(* Logix 5000 project; controller PLC_MCC1300_75F1 vendor 1 type 14 code 166 rev 32.11; software revision 32.04; part 55 of 83 *)
(* tags used below, declared in another part *)
   CM_AreaStackerToLine_JS1 : CM_AreaStackerToLine;
   CM_AreaStackerToLine_JS1_Sync : CM_AreaStackerToLine;
   CM_ConveyorStackerToLine_JS1_Sync : CM_ConveyorStackerToLine;
   Convoy_SL_DATA_NULL : UDT_Convoy_SL;
   GP_AccessArea_M311S_STC : GP_AccessArea_STC;
   GP_InvertCapxLite : GP_InvertCapxLite;
   GP_M311A : GP_Rotator;
   GP_OB_InitializeMain : GP_OB_Initialize;
   GP_ScadaPlate : GP_ScadaPlate;
   Gp_SpaceConvUtilities_V1 : GP_SpaceConvUtilities_V1;
   M310B : MAC_Conveyor;
   M310B_Data : UDT_Convoy_SL;
   M310B_SpaceConv_Utilities : SpaceConv_Utilities;
   M311 : MAC_Conveyor;
   M311_ALM : MAC_Conveyor_ALM;
   M311_Data : UDT_Convoy_SL;
   M311_dLastRotationA_ID : DINT;
   M311_HMR : MAC_Conveyor_HMR;
   M311_HMW : MAC_Conveyor_HMW;
   M311_M1_DR : AXIS_CIP_DRIVE;
   M311_M1_DR_IN_MAM : MOTION_INSTRUCTION;
   M311_SpaceConv_Utilities : SpaceConv_Utilities;
   M311_TON_Synchro_timeout : TIMER;
   M311_xOS_SentToCullet : BOOL;
   M311_xSendCulletReqActive : BOOL;
   M311_xSensorTimeout : BOOL;
   M311A : MAC_Rotator;
   M311A_Data : UDT_Convoy_SL;
   M311A_HMR : MAC_Rotator_HMR;
   M311A_HMW : MAC_Rotator_HMW;
   M311A_M1_DR : AXIS_CIP_DRIVE;
   M311A_M1_DR_IN_MAM : MOTION_INSTRUCTION;
   M311A_rLastPosition : REAL;
   M311M312_OffsetBaricentre_cmm : DINT;
   M312 : MAC_Conveyor_Single;
   M312_Data : UDT_Convoy_SL;
   M312_SpaceConv_Utilities : SpaceConv_Utilities;
   O : INT[128];
   Sbr_OUT_ReqRot_CW : BOOL;
   TMP_d : DINT;
   TMP_dActualOnLHS : DINT;
   TMP_dDecelerationPositionEndConveyor : DINT;
   TMP_dMissingOnLHS : DINT;
   TMP_dOffsetLoadUnload_cmm : DINT;
   TMP_HeadPos : DINT;
   TMP_Portrait : BOOL;
   TMP_SendToCullet : BOOL;
   TMP_x : BOOL;
   TMP_xConveyorOfStartCleaning : BOOL;
   TMP_xEnableZoneCleaning : BOOL;
   TMP_xJustOnePlateMissing : BOOL;
   TMP_xLiteThisDestPresent : BOOL;
   x311PortraitMode : BOOL;
   xAlwaysOFF : BOOL;
   xAlwaysON : BOOL;
   xDebugOFF : BOOL;
   Z401 : MAC_Zone;
   Z401_HMI_rgtPlateScada_Internal : HMI_LiteData[5,2,7];
   Z401_HMR : MAC_Zone_HMR;
   Z401S_INPUT_xSafetyAreaPopup : BOOL;
(* MainProgram, continued *)

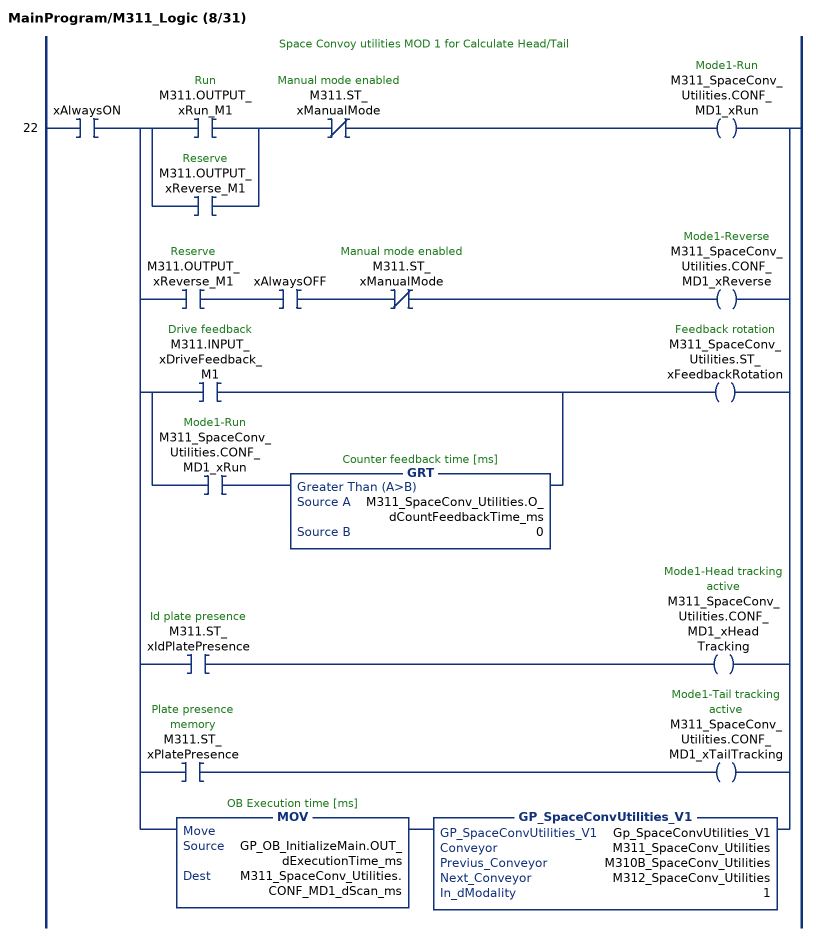
   [picture p890: MainProgram/M311_Logic rungs 22-22]
   // Space Convoy utilities MOD 1 for Calculate Head/Tail
   22: XIC(xAlwaysON)[[XIC(M311.OUTPUT_xRun_M1) ,XIC(M311.OUTPUT_xReverse_M1) ] XIO(M311.ST_xManualMode) OTE(M311_SpaceConv_Utilities.CONF_MD1_xRun) ,XIC(M311.OUTPUT_xReverse_M1) XIC(xAlwaysOFF) XIO(M311.ST_xManualMode) OTE(M311_SpaceConv_Utilities.CONF_MD1_xReverse) ,[XIC(M311.INPUT_xDriveFeedback_M1) ,XIC(M311_SpaceConv_Utilities.CONF_MD1_xRun) GRT(M311_SpaceConv_Utilities.O_dCountFeedbackTime_ms,0) ] OTE(M311_SpaceConv_Utilities.ST_xFeedbackRotation) ,XIC(M311.ST_xIdPlatePresence) OTE(M311_SpaceConv_Utilities.CONF_MD1_xHeadTracking) ,XIC(M311.ST_xPlatePresence) OTE(M311_SpaceConv_Utilities.CONF_MD1_xTailTracking) ,MOV(GP_OB_InitializeMain.OUT_dExecutionTime_ms,M311_SpaceConv_Utilities.CONF_MD1_dScan_ms) GP_SpaceConvUtilities_V1(Gp_SpaceConvUtilities_V1,M311_SpaceConv_Utilities,M310B_SpaceConv_Utilities,M312_SpaceConv_Utilities,1) ];
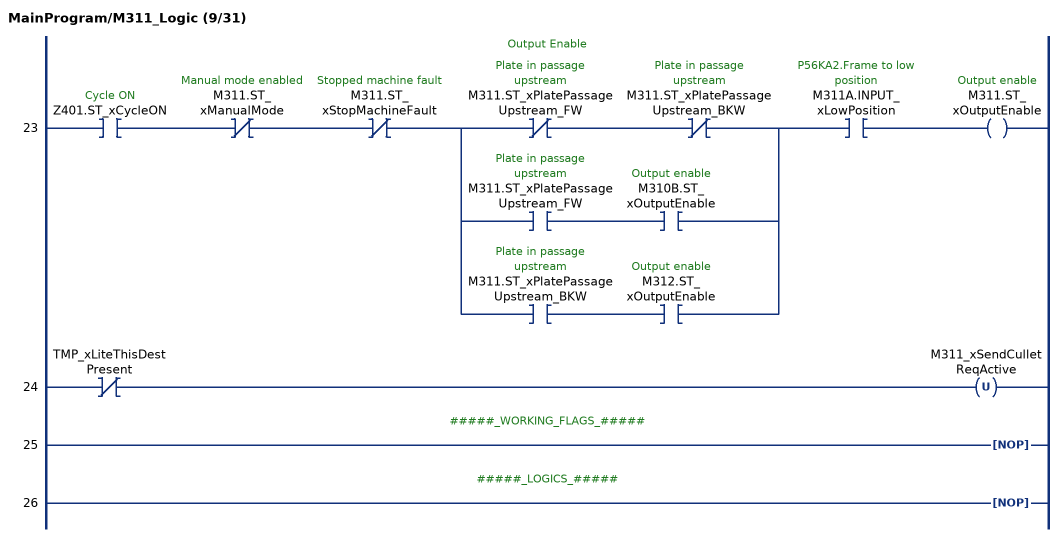
   // Output Enable
   23: XIC(Z401.ST_xCycleON)XIO(M311.ST_xManualMode)XIO(M311.ST_xStopMachineFault)[XIO(M311.ST_xPlatePassageUpstream_FW) XIO(M311.ST_xPlatePassageUpstream_BKW) ,XIC(M311.ST_xPlatePassageUpstream_FW) XIC(M310B.ST_xOutputEnable) ,XIC(M311.ST_xPlatePassageUpstream_BKW) XIC(M312.ST_xOutputEnable) ]XIC(M311A.INPUT_xLowPosition)OTE(M311.ST_xOutputEnable);
   24: XIO(TMP_xLiteThisDestPresent)OTU(M311_xSendCulletReqActive);
   // #####_WORKING_FLAGS_#####
   25: NOP();
   // #####_LOGICS_#####
   26: NOP();
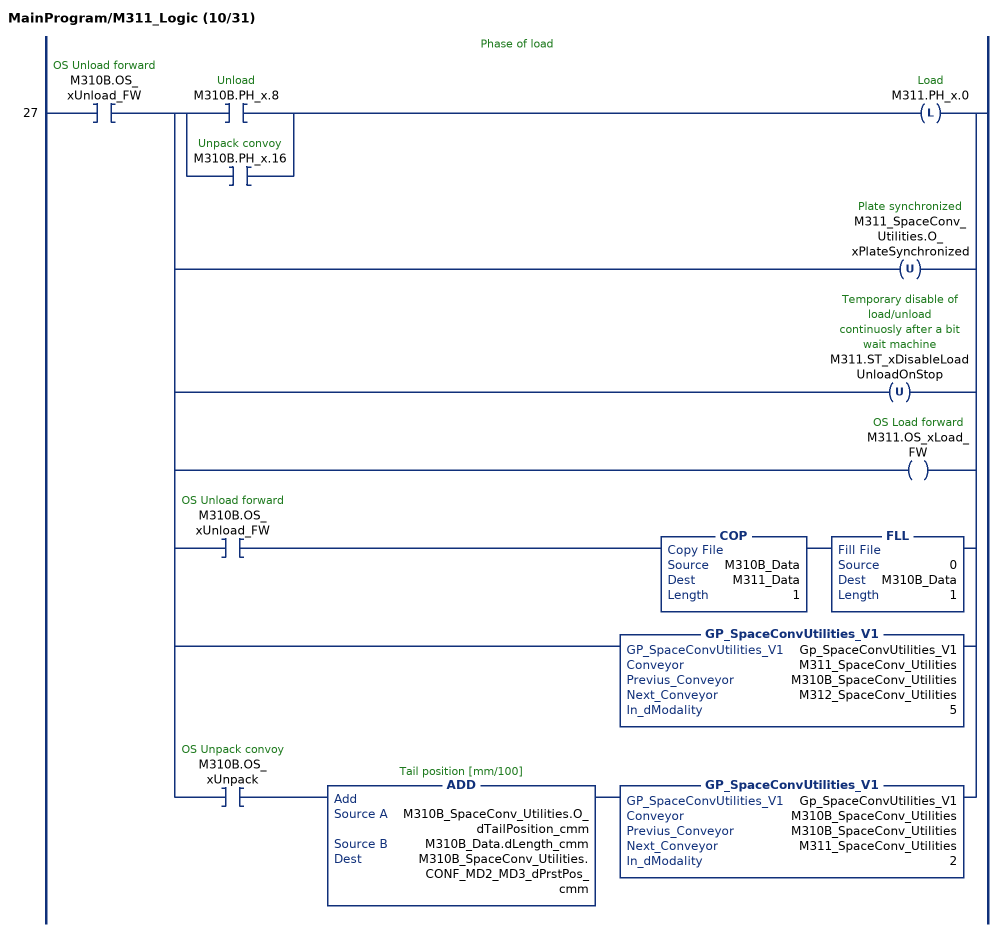
   // Phase of load
   27: XIC(M310B.OS_xUnload_FW)[[XIC(M310B.PH_x.8) ,XIC(M310B.PH_x.16) ] OTL(M311.PH_x.0) ,OTU(M311_SpaceConv_Utilities.O_xPlateSynchronized) ,OTU(M311.ST_xDisableLoadUnloadOnStop) ,OTE(M311.OS_xLoad_FW) ,XIC(M310B.OS_xUnload_FW) COP(M310B_Data,M311_Data,1) FLL(0,M310B_Data,1) ,GP_SpaceConvUtilities_V1(Gp_SpaceConvUtilities_V1,M311_SpaceConv_Utilities,M310B_SpaceConv_Utilities,M312_SpaceConv_Utilities,5) ,XIC(M310B.OS_xUnpack) ADD(M310B_SpaceConv_Utilities.O_dTailPosition_cmm,M310B_Data.dLength_cmm,M310B_SpaceConv_Utilities.CONF_MD2_MD3_dPrstPos_cmm) GP_SpaceConvUtilities_V1(Gp_SpaceConvUtilities_V1,M310B_SpaceConv_Utilities,M310B_SpaceConv_Utilities,M311_SpaceConv_Utilities,2) ];
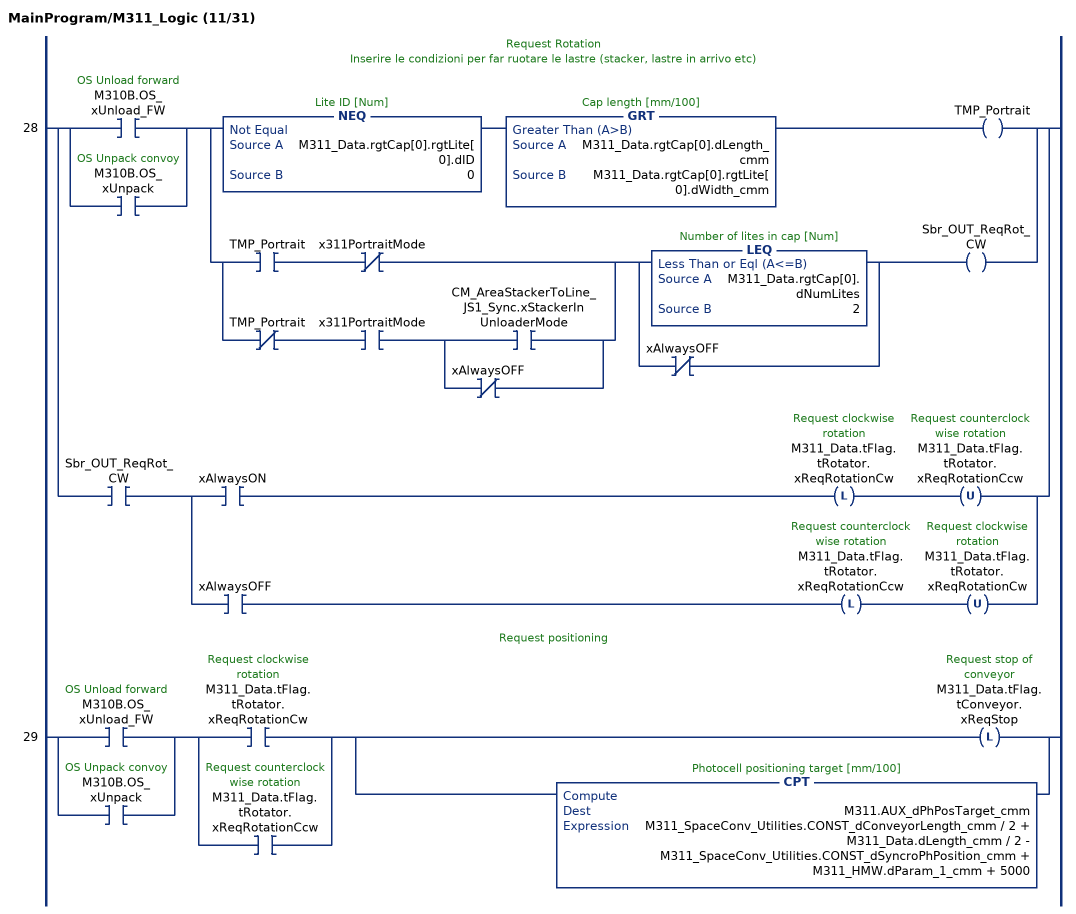
   // Request Rotation
   // Inserire le condizioni per far ruotare le lastre (stacker, lastre in arrivo etc)
   28: [[XIC(M310B.OS_xUnload_FW) ,XIC(M310B.OS_xUnpack) ] [NEQ(M311_Data.rgtCap[0].rgtLite[0].dID,0) GRT(M311_Data.rgtCap[0].dLength_cmm,M311_Data.rgtCap[0].rgtLite[0].dWidth_cmm) OTE(TMP_Portrait) ,[XIC(TMP_Portrait) XIO(x311PortraitMode) ,XIO(TMP_Portrait) XIC(x311PortraitMode) [XIC(CM_AreaStackerToLine_JS1_Sync.xStackerInUnloaderMode) ,XIO(xAlwaysOFF) ] ] [LEQ(M311_Data.rgtCap[0].dNumLites,2) ,XIO(xAlwaysOFF) ] OTE(Sbr_OUT_ReqRot_CW) ] ,XIC(Sbr_OUT_ReqRot_CW) [XIC(xAlwaysON) OTL(M311_Data.tFlag.tRotator.xReqRotationCw) OTU(M311_Data.tFlag.tRotator.xReqRotationCcw) ,XIC(xAlwaysOFF) OTL(M311_Data.tFlag.tRotator.xReqRotationCcw) OTU(M311_Data.tFlag.tRotator.xReqRotationCw) ] ];
   // Request positioning
   29: [XIC(M310B.OS_xUnload_FW) ,XIC(M310B.OS_xUnpack) ][XIC(M311_Data.tFlag.tRotator.xReqRotationCw) ,XIC(M311_Data.tFlag.tRotator.xReqRotationCcw) ][OTL(M311_Data.tFlag.tConveyor.xReqStop) ,CPT(M311.AUX_dPhPosTarget_cmm,M311_SpaceConv_Utilities.CONST_dConveyorLength_cmm / 2 + M311_Data.dLength_cmm / 2 - M311_SpaceConv_Utilities.CONST_dSyncroPhPosition_cmm + M311_HMW.dParam_1_cmm + 5000) ];
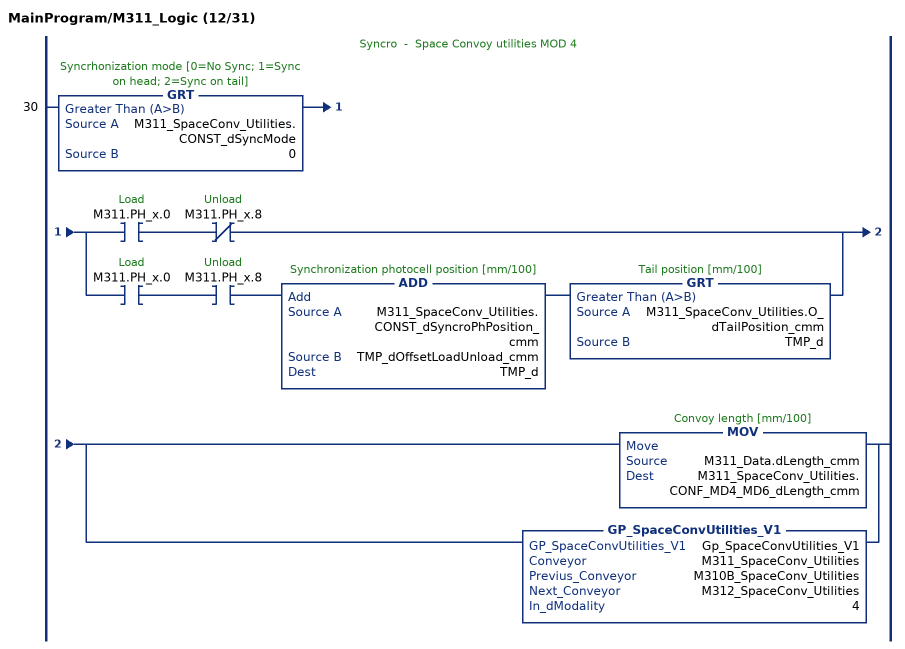
   // Syncro  -  Space Convoy utilities MOD 4
   30: GRT(M311_SpaceConv_Utilities.CONST_dSyncMode,0)[XIC(M311.PH_x.0) XIO(M311.PH_x.8) ,XIC(M311.PH_x.0) XIC(M311.PH_x.8) ADD(M311_SpaceConv_Utilities.CONST_dSyncroPhPosition_cmm,TMP_dOffsetLoadUnload_cmm,TMP_d) GRT(M311_SpaceConv_Utilities.O_dTailPosition_cmm,TMP_d) ][MOV(M311_Data.dLength_cmm,M311_SpaceConv_Utilities.CONF_MD4_MD6_dLength_cmm) ,GP_SpaceConvUtilities_V1(Gp_SpaceConvUtilities_V1,M311_SpaceConv_Utilities,M310B_SpaceConv_Utilities,M312_SpaceConv_Utilities,4) ];
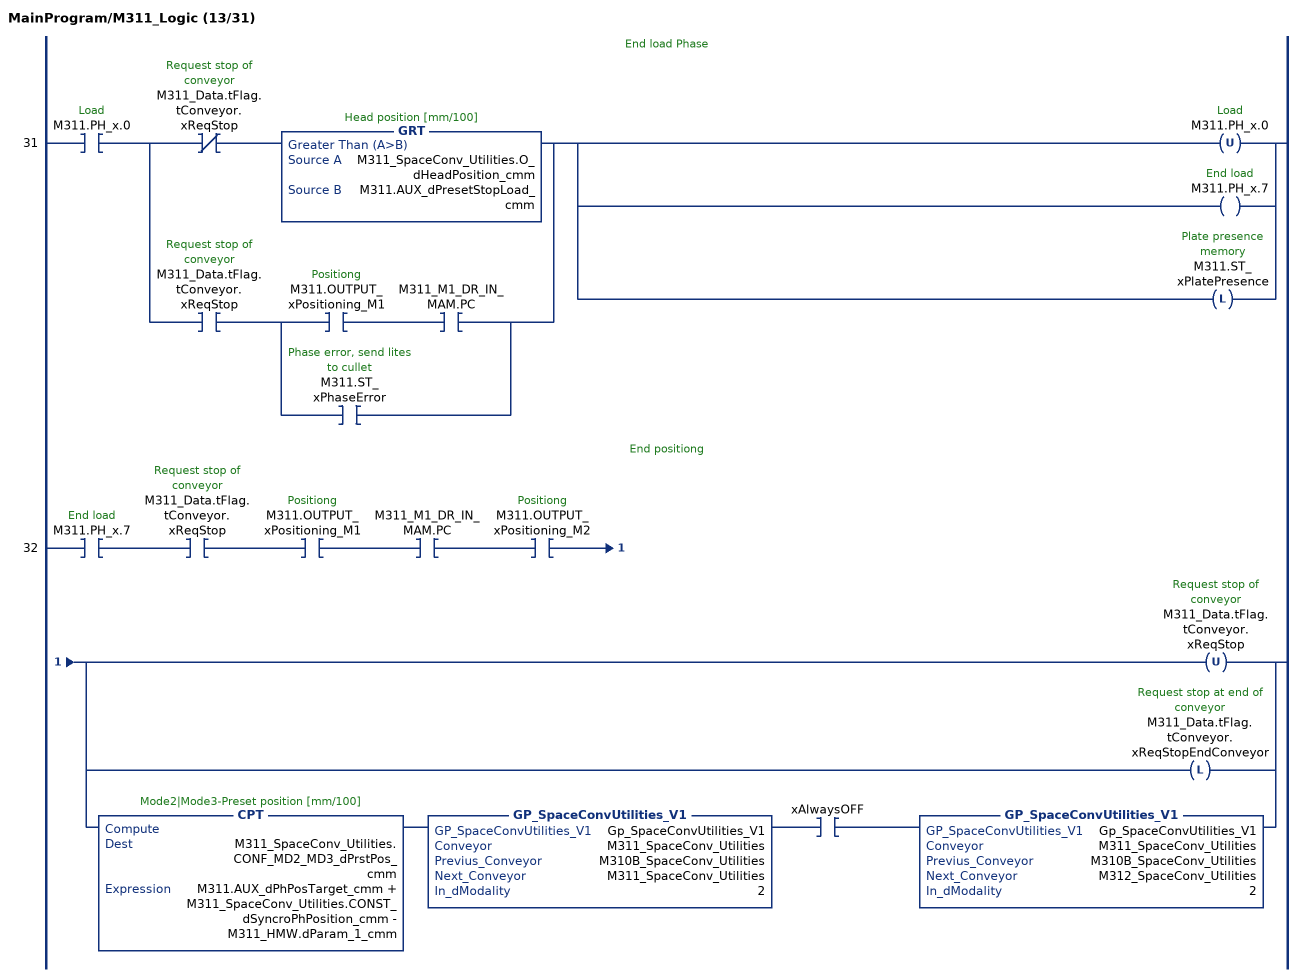
   // End load Phase
   31: XIC(M311.PH_x.0)[XIO(M311_Data.tFlag.tConveyor.xReqStop) GRT(M311_SpaceConv_Utilities.O_dHeadPosition_cmm,M311.AUX_dPresetStopLoad_cmm) ,XIC(M311_Data.tFlag.tConveyor.xReqStop) [XIC(M311.OUTPUT_xPositioning_M1) XIC(M311_M1_DR_IN_MAM.PC) ,XIC(M311.ST_xPhaseError) ] ][OTU(M311.PH_x.0) ,OTE(M311.PH_x.7) ,OTL(M311.ST_xPlatePresence) ];
   // End positiong
   32: XIC(M311.PH_x.7)XIC(M311_Data.tFlag.tConveyor.xReqStop)XIC(M311.OUTPUT_xPositioning_M1)XIC(M311_M1_DR_IN_MAM.PC)XIC(M311.OUTPUT_xPositioning_M2)[OTU(M311_Data.tFlag.tConveyor.xReqStop) ,OTL(M311_Data.tFlag.tConveyor.xReqStopEndConveyor) ,CPT(M311_SpaceConv_Utilities.CONF_MD2_MD3_dPrstPos_cmm,M311.AUX_dPhPosTarget_cmm + M311_SpaceConv_Utilities.CONST_dSyncroPhPosition_cmm - M311_HMW.dParam_1_cmm) GP_SpaceConvUtilities_V1(Gp_SpaceConvUtilities_V1,M311_SpaceConv_Utilities,M310B_SpaceConv_Utilities,M311_SpaceConv_Utilities,2) XIC(xAlwaysOFF) GP_SpaceConvUtilities_V1(Gp_SpaceConvUtilities_V1,M311_SpaceConv_Utilities,M310B_SpaceConv_Utilities,M312_SpaceConv_Utilities,2) ];
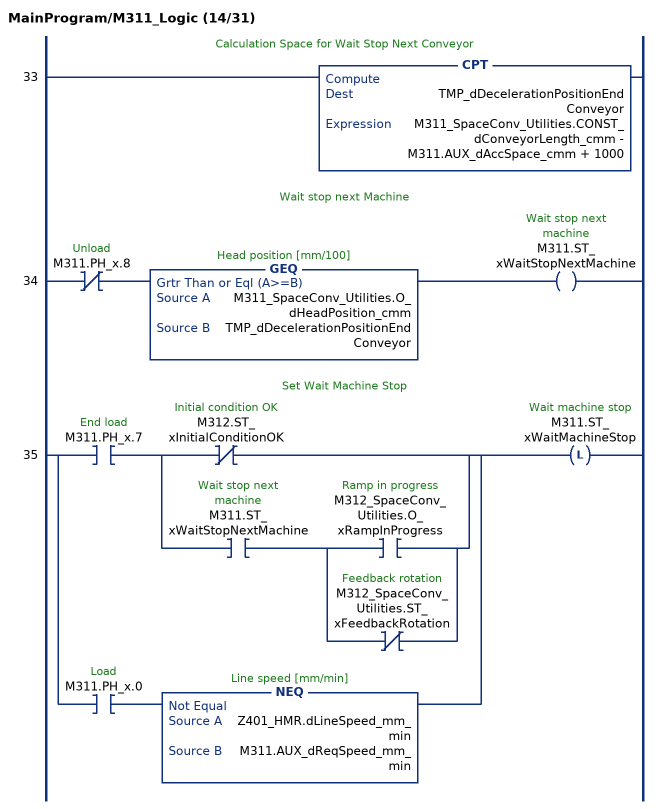
   // Calculation Space for Wait Stop Next Conveyor
   33: CPT(TMP_dDecelerationPositionEndConveyor,M311_SpaceConv_Utilities.CONST_dConveyorLength_cmm - M311.AUX_dAccSpace_cmm + 1000);
   // Wait stop next Machine
   34: XIO(M311.PH_x.8)GEQ(M311_SpaceConv_Utilities.O_dHeadPosition_cmm,TMP_dDecelerationPositionEndConveyor)OTE(M311.ST_xWaitStopNextMachine);
   // Set Wait Machine Stop
   35: [XIC(M311.PH_x.7) [XIO(M312.ST_xInitialConditionOK) ,XIC(M311.ST_xWaitStopNextMachine) [XIC(M312_SpaceConv_Utilities.O_xRampInProgress) ,XIO(M312_SpaceConv_Utilities.ST_xFeedbackRotation) ] ] ,XIC(M311.PH_x.0) NEQ(Z401_HMR.dLineSpeed_mm_min,M311.AUX_dReqSpeed_mm_min) ]OTL(M311.ST_xWaitMachineStop);
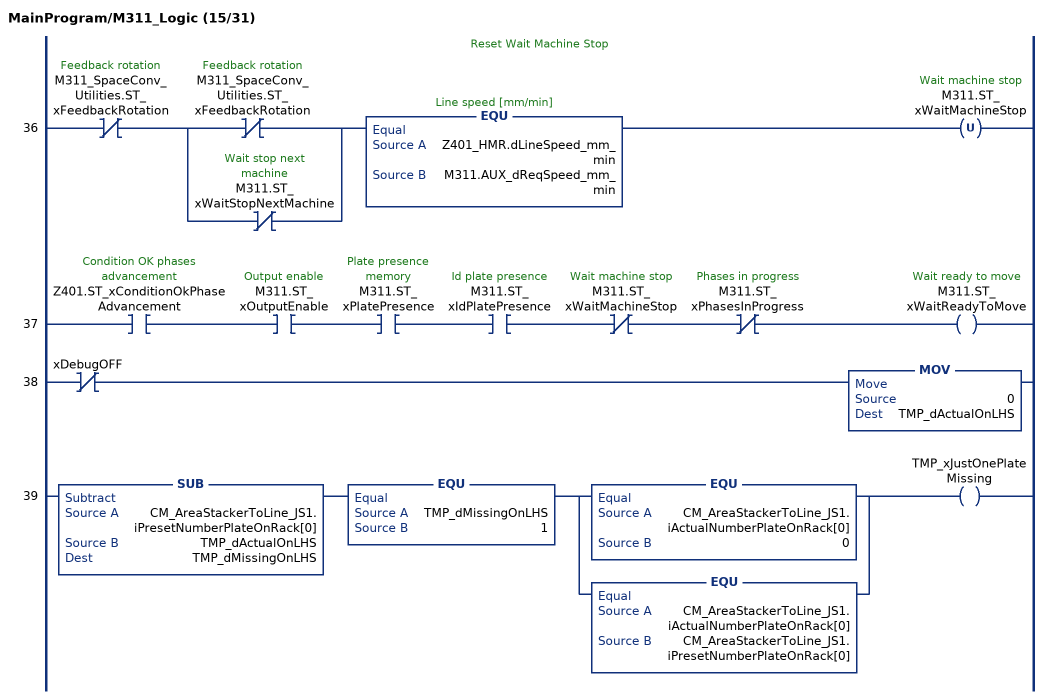
   // Reset Wait Machine Stop
   36: XIO(M311_SpaceConv_Utilities.ST_xFeedbackRotation)[XIO(M311_SpaceConv_Utilities.ST_xFeedbackRotation) ,XIO(M311.ST_xWaitStopNextMachine) ]EQU(Z401_HMR.dLineSpeed_mm_min,M311.AUX_dReqSpeed_mm_min)OTU(M311.ST_xWaitMachineStop);
   37: XIC(Z401.ST_xConditionOkPhaseAdvancement)XIC(M311.ST_xOutputEnable)XIC(M311.ST_xPlatePresence)XIC(M311.ST_xIdPlatePresence)XIO(M311.ST_xWaitMachineStop)XIO(M311.ST_xPhasesInProgress)OTE(M311.ST_xWaitReadyToMove);
   38: XIO(xDebugOFF)MOV(0,TMP_dActualOnLHS);
   39: SUB(CM_AreaStackerToLine_JS1.iPresetNumberPlateOnRack[0],TMP_dActualOnLHS,TMP_dMissingOnLHS)EQU(TMP_dMissingOnLHS,1)[EQU(CM_AreaStackerToLine_JS1.iActualNumberPlateOnRack[0],0) ,EQU(CM_AreaStackerToLine_JS1.iActualNumberPlateOnRack[0],CM_AreaStackerToLine_JS1.iPresetNumberPlateOnRack[0]) ]OTE(TMP_xJustOnePlateMissing);
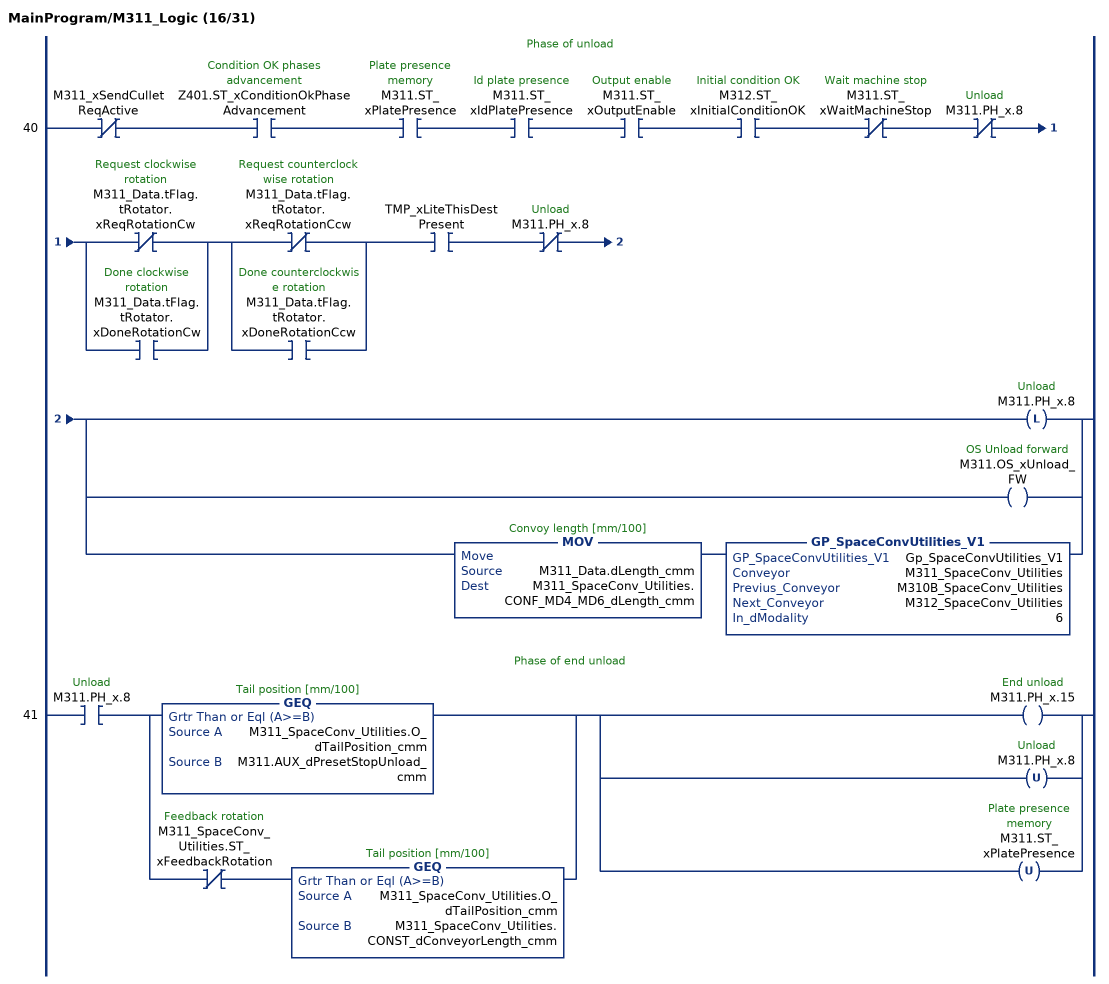
   // Phase of unload
   40: XIO(M311_xSendCulletReqActive)XIC(Z401.ST_xConditionOkPhaseAdvancement)XIC(M311.ST_xPlatePresence)XIC(M311.ST_xIdPlatePresence)XIC(M311.ST_xOutputEnable)XIC(M312.ST_xInitialConditionOK)XIO(M311.ST_xWaitMachineStop)XIO(M311.PH_x.8)[XIO(M311_Data.tFlag.tRotator.xReqRotationCw) ,XIC(M311_Data.tFlag.tRotator.xDoneRotationCw) ][XIO(M311_Data.tFlag.tRotator.xReqRotationCcw) ,XIC(M311_Data.tFlag.tRotator.xDoneRotationCcw) ]XIC(TMP_xLiteThisDestPresent)XIO(M311.PH_x.8)[OTL(M311.PH_x.8) ,OTE(M311.OS_xUnload_FW) ,MOV(M311_Data.dLength_cmm,M311_SpaceConv_Utilities.CONF_MD4_MD6_dLength_cmm) GP_SpaceConvUtilities_V1(Gp_SpaceConvUtilities_V1,M311_SpaceConv_Utilities,M310B_SpaceConv_Utilities,M312_SpaceConv_Utilities,6) ];
   // Phase of end unload
   41: XIC(M311.PH_x.8)[GEQ(M311_SpaceConv_Utilities.O_dTailPosition_cmm,M311.AUX_dPresetStopUnload_cmm) ,XIO(M311_SpaceConv_Utilities.ST_xFeedbackRotation) GEQ(M311_SpaceConv_Utilities.O_dTailPosition_cmm,M311_SpaceConv_Utilities.CONST_dConveyorLength_cmm) ][OTE(M311.PH_x.15) ,OTU(M311.PH_x.8) ,OTU(M311.ST_xPlatePresence) ];
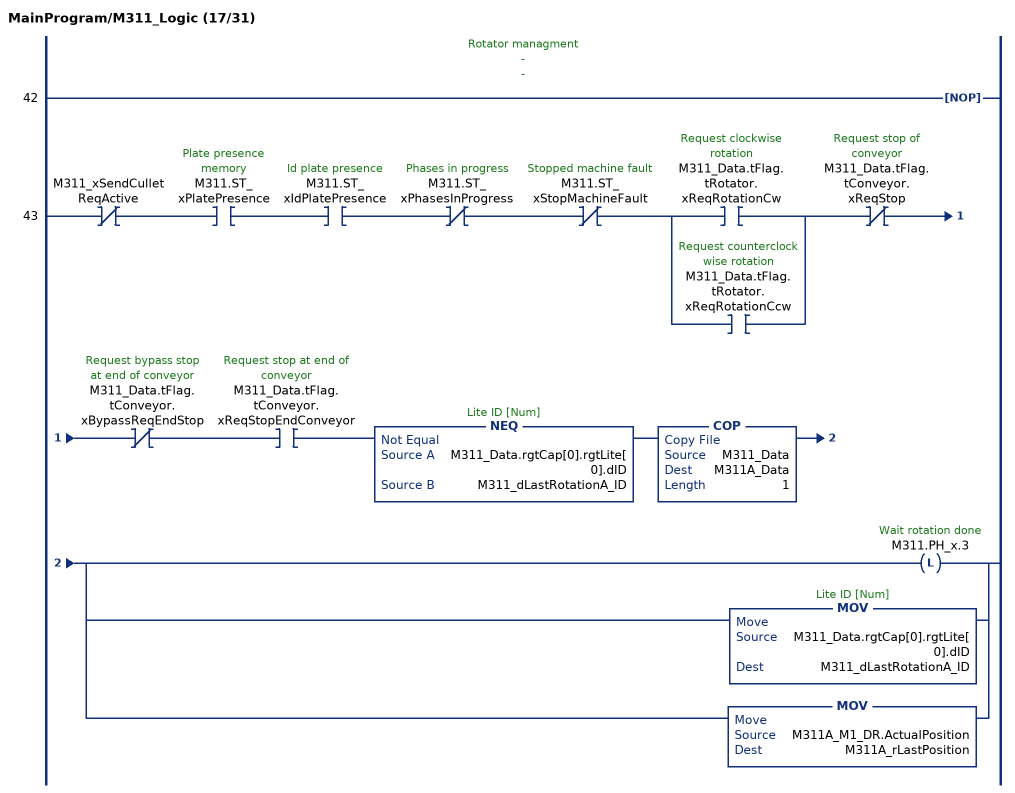
   // Rotator managment
   // -
   // -
   42: NOP();
   43: XIO(M311_xSendCulletReqActive)XIC(M311.ST_xPlatePresence)XIC(M311.ST_xIdPlatePresence)XIO(M311.ST_xPhasesInProgress)XIO(M311.ST_xStopMachineFault)[XIC(M311_Data.tFlag.tRotator.xReqRotationCw) ,XIC(M311_Data.tFlag.tRotator.xReqRotationCcw) ]XIO(M311_Data.tFlag.tConveyor.xReqStop)XIO(M311_Data.tFlag.tConveyor.xBypassReqEndStop)XIC(M311_Data.tFlag.tConveyor.xReqStopEndConveyor)NEQ(M311_Data.rgtCap[0].rgtLite[0].dID,M311_dLastRotationA_ID)COP(M311_Data,M311A_Data,1)[OTL(M311.PH_x.3) ,MOV(M311_Data.rgtCap[0].rgtLite[0].dID,M311_dLastRotationA_ID) ,MOV(M311A_M1_DR.ActualPosition,M311A_rLastPosition) ];